   "Carrier_69_SpareSafetyInput(2_6)" AT %I3814.6 : Bool;   // SPARE SAFETY INPUT
   "Carrier_69_SpareSafetyInput(2_7)" AT %I3814.7 : Bool;   // SPARE SAFETY INPUT
   "Carrier_69_Slot3_SafetyOutput" AT %IW3815 : Word;   // SLOT 3 SAFETY OUTPUT WORD
   "Carrier_69_Crash_Detect_OK" AT %I3815.0 : Bool;   // CARRIER CRASH DETECT
   "Carrier_69_SpareSafetyOutput(3_1)" AT %I3815.1 : Bool;   // SPARE SAFETY OUTPUT
   "Carrier_69_SpareSafetyOutput(3_2)" AT %I3815.2 : Bool;   // SPARE SAFETY OUTPUT
   "Carrier_69_SpareSafetyOutput(3_3)" AT %I3815.3 : Bool;   // SPARE SAFETY OUTPUT
   "Carrier_69_SpareSafetyOutput(3_4)" AT %I3815.4 : Bool;   // SPARE SAFETY OUTPUT
   "Carrier_69_SpareSafetyOutput(3_5)" AT %I3815.5 : Bool;   // SPARE SAFETY OUTPUT
   "Carrier_69_SpareSafetyOutput(3_6)" AT %I3815.6 : Bool;   // SPARE SAFETY OUTPUT
   "Carrier_69_SpareSafetyOutput(3_7)" AT %I3815.7 : Bool;   // SPARE SAFETY OUTPUT
   "Carrier_69_Slot4_Input" AT %IW3816 : Word;   // SLOT 4 INPUT WORD
   "Carrier_69_480VPowerOn_MDCB1" AT %I3816.0 : Bool;   // 480 VAC POWER ON MDCB 1
   "Carrier_69_SpareInput(4_1)" AT %I3816.1 : Bool;   // SPARE INPUT
   "Carrier_69_SpareInput(4_2)" AT %I3816.2 : Bool;   // SPARE INPUT
   "Carrier_69_SitopSelectStatus" AT %I3816.3 : Bool;   // SITOP SELECT STATUS
   "Carrier_69_DCsupplyOnPSCB2" AT %I3816.4 : Bool;   // DC SUPPLY ON PSCB 2
   "Carrier_69_SpareInput(4_5)" AT %I3816.5 : Bool;   // SPARE INPUT
   "Carrier_69_SpareInput(4_6)" AT %I3816.6 : Bool;   // SPARE INPUT
   "Carrier_69_SpareInput(4_7)" AT %I3816.7 : Bool;   // SPARE INPUT
   "Carrier_69_PB1_ProdHoldLH" AT %I3817.0 : Bool;   // PB 1 PRODUCTION HOLD LH
   "Carrier_69_PB2_ResetLH" AT %I3817.1 : Bool;   // PB 2 RESET LH
   "Carrier_69_PB3_ProdHoldRH" AT %I3817.2 : Bool;   // PB 3 PRODUCTION HOLD RH
   "Carrier_69_PB4_ResetRH" AT %I3817.3 : Bool;   // PB 4 RESET RH
   "Carrier_69_SpareInput(4_14)" AT %I3817.4 : Bool;   // SPARE INPUT
   "Carrier_69_SpareInput(4_15)" AT %I3817.5 : Bool;   // SPARE INPUT
   "Carrier_69_SpareInput(4_16)" AT %I3817.6 : Bool;   // SPARE INPUT
   "Carrier_69_SpareInput(4_17)" AT %I3817.7 : Bool;   // SPARE INPUT
   "Carrier_69_Slot5_Output" AT %IW3818 : Word;   // SLOT 5 OUTPUT WORD
   "Carrier_69_IRD400_HMI_24VDC_ENABLE" AT %I3818.0 : Bool;   // IRD 400 PANEL HMI 24V DC POWER
   "Carrier_69_FaultLight_LH" AT %I3818.1 : Bool;   // FAULT LIGHT LH
   "Carrier_69_RunLight_LH" AT %I3818.2 : Bool;   // RUN LIGHT LH
   "Carrier_69_FaultLight_RH" AT %I3818.3 : Bool;   // FAULT LIGHT RH
   "Carrier_69_RunLight_RH" AT %I3818.4 : Bool;   // RUN LIGHT RH
   "Carrier_69_SpareOutput(5_5)" AT %I3818.5 : Bool;   // SPARE OUTPUT
   "Carrier_69_SpareOutput(5_6)" AT %I3818.6 : Bool;   // SPARE OUTPUT
   "Carrier_69_SpareOutput(5_7)" AT %I3818.7 : Bool;   // SPARE OUTPUT
   "Carrier_69_ActualSpeed" AT %IW3820 : Word;   // ACTUAL SPEED
   "Carrier_69_CarrierDriveAlarm" AT %IW3822 : Word;   // CARRIER DRIVE ALARM
   "Carrier_69_CarrierDriveWarning" AT %IW3824 : Word;   // CARRIER DRIVE WARNING
   "Carrier_70_Status" AT %IW3850 : Word;   // CARRIER STATUS WORD
   "Carrier_70_Status.0" AT %I3850.0 : Bool;   // HEARTBEAT
   "Carrier_70_Status.1" AT %I3850.1 : Bool;   // MANUAL
   "Carrier_70_Status.2" AT %I3850.2 : Bool;   // IN_AUTO
   "Carrier_70_Status.3" AT %I3850.3 : Bool;   // POSITIONING_COMPLETE
   "Carrier_70_Status.4" AT %I3850.4 : Bool;   // PRODUCTION HOLD
   "Carrier_70_Status.5" AT %I3850.5 : Bool;   // CARRIER MOVING FORWARD
   "Carrier_70_Status.6" AT %I3850.6 : Bool;   // CARRIER MOVING REVERSE
   "Carrier_70_Status.7" AT %I3850.7 : Bool;   // CARRIER FAULT
   "Carrier_70_Status.8" AT %I3851.0 : Bool;   // CRASH DETECT TRIPPED
   "Carrier_70_Status.9" AT %I3851.1 : Bool;
   "Carrier_70_Status.10" AT %I3851.2 : Bool;
   "Carrier_70_Status.11" AT %I3851.3 : Bool;
   "Carrier_70_Status.12" AT %I3851.4 : Bool;
   "Carrier_70_Status.13" AT %I3851.5 : Bool;
   "Carrier_70_Status.14" AT %I3851.6 : Bool;
   "Carrier_70_Status.15" AT %I3851.7 : Bool;
   "Carrier_70_SDCFaultCode" AT %IW3852 : Word;   // SDC FAULT CODE
   "Carrier_70_CarrierPosition" AT %ID3854 : DWord;   // CARRIER POSITION
   "Carrier_70_CarrierNumber" AT %IW3858 : Word;   // CARRIER NUMBER
   "Carrier_70_G120DControlWord" AT %IW3860 : Word;   // G120D_STW1_CONTROL
   "Carrier_70_G120DControlWord.0" AT %I3860.0 : Bool;   // Bit_00_ON
   "Carrier_70_G120DControlWord.1" AT %I3860.1 : Bool;   // Bit_01_AUS2_INH
   "Carrier_70_G120DControlWord.2" AT %I3860.2 : Bool;   // Bit_02_AUS3_STOP
   "Carrier_70_G120DControlWord.3" AT %I3860.3 : Bool;   // Bit_03_EN
   "Carrier_70_G120DControlWord.4" AT %I3860.4 : Bool;   // Bit_04_EN_RAMP
   "Carrier_70_G120DControlWord.5" AT %I3860.5 : Bool;   // Bit_05_START_RAMP
   "Carrier_70_G120DControlWord.6" AT %I3860.6 : Bool;   // Bit_06_SETPOINT
   "Carrier_70_G120DControlWord.7" AT %I3860.7 : Bool;   // Bit_07_RESET
   "Carrier_70_G120DControlWord.8" AT %I3861.0 : Bool;   // Bit_08_JOG_R
   "Carrier_70_G120DControlWord.9" AT %I3861.1 : Bool;   // Bit_09_JOG_L
   "Carrier_70_G120DControlWord.10" AT %I3861.2 : Bool;   // Bit_10_CONTR_PLC
   "Carrier_70_G120DControlWord.11" AT %I3861.3 : Bool;   // Bit_11_REVERSE
   "Carrier_70_G120DControlWord.12" AT %I3861.4 : Bool;   // Bit_12_BRAKE_RELEASE
   "Carrier_70_G120DControlWord.13" AT %I3861.5 : Bool;   // Bit_13_DDS
   "Carrier_70_G120DControlWord.14" AT %I3861.6 : Bool;   // Bit_14_DO0
   "Carrier_70_G120DControlWord.15" AT %I3861.7 : Bool;   // Bit_15_DO1
   "Carrier_70_G120DStatusWord" AT %IW3862 : Word;   // G120D_ZSW1_STATUS
   "Carrier_70_G120DStatusWord.0" AT %I3862.0 : Bool;   // Bit_00_READY_RUN
   "Carrier_70_G120DStatusWord.1" AT %I3862.1 : Bool;   // Bit_01_READY_ON
   "Carrier_70_G120DStatusWord.2" AT %I3862.2 : Bool;   // Bit_02_ENABLE
   "Carrier_70_G120DStatusWord.3" AT %I3862.3 : Bool;   // Bit_03_FAULT
   "Carrier_70_G120DStatusWord.4" AT %I3862.4 : Bool;   // Bit_04_OFF2
   "Carrier_70_G120DStatusWord.5" AT %I3862.5 : Bool;   // Bit_05_OFF3
   "Carrier_70_G120DStatusWord.6" AT %I3862.6 : Bool;   // Bit_06_LOCK_OUT
   "Carrier_70_G120DStatusWord.7" AT %I3862.7 : Bool;   // Bit_07_WARN
   "Carrier_70_G120DStatusWord.8" AT %I3863.0 : Bool;   // Bit_08_NO_DEVIATION
   "Carrier_70_G120DStatusWord.9" AT %I3863.1 : Bool;   // Bit_09_CONTR_PLC
   "Carrier_70_G120DStatusWord.10" AT %I3863.2 : Bool;   // Bit_10_F_MAX
   "Carrier_70_G120DStatusWord.11" AT %I3863.3 : Bool;   // Bit_11_LIMIT_REACHED
   "Carrier_70_G120DStatusWord.12" AT %I3863.4 : Bool;   // Bit_12_BRAKE_OPEN
   "Carrier_70_G120DStatusWord.13" AT %I3863.5 : Bool;   // Bit_13_NO_OVERTEMP
   "Carrier_70_G120DStatusWord.14" AT %I3863.6 : Bool;   // Bit_14_CW_CCW
   "Carrier_70_G120DStatusWord.15" AT %I3863.7 : Bool;   // Bit_15_OVERL
   "Carrier_70_Slot2_Input" AT %IW3864 : Word;   // SLOT 2 INPUT WORD
   "Carrier_70_CrashDetectSW" AT %I3864.0 : Bool;   // CRASH DETECT SW
   "Carrier_70_SpareSafetyInput(2_1)" AT %I3864.1 : Bool;   // SPARE SAFETY INPUT
   "Carrier_70_SpareSafetyInput(2_2)" AT %I3864.2 : Bool;   // SPARE SAFETY INPUT
   "Carrier_70_SpareSafetyInput(2_3)" AT %I3864.3 : Bool;   // SPARE SAFETY INPUT
   "Carrier_70_SpareSafetyInput(2_4)" AT %I3864.4 : Bool;   // SPARE SAFETY INPUT
   "Carrier_70_SpareSafetyInput(2_5)" AT %I3864.5 : Bool;   // SPARE SAFETY INPUT
   "Carrier_70_SpareSafetyInput(2_6)" AT %I3864.6 : Bool;   // SPARE SAFETY INPUT
   "Carrier_70_SpareSafetyInput(2_7)" AT %I3864.7 : Bool;   // SPARE SAFETY INPUT
   "Carrier_70_Slot3_SafetyOutput" AT %IW3865 : Word;   // SLOT 3 SAFETY OUTPUT WORD
   "Carrier_70_Crash_Detect_OK" AT %I3865.0 : Bool;   // CARRIER CRASH DETECT
   "Carrier_70_SpareSafetyOutput(3_1)" AT %I3865.1 : Bool;   // SPARE SAFETY OUTPUT
   "Carrier_70_SpareSafetyOutput(3_2)" AT %I3865.2 : Bool;   // SPARE SAFETY OUTPUT
   "Carrier_70_SpareSafetyOutput(3_3)" AT %I3865.3 : Bool;   // SPARE SAFETY OUTPUT
   "Carrier_70_SpareSafetyOutput(3_4)" AT %I3865.4 : Bool;   // SPARE SAFETY OUTPUT
   "Carrier_70_SpareSafetyOutput(3_5)" AT %I3865.5 : Bool;   // SPARE SAFETY OUTPUT
   "Carrier_70_SpareSafetyOutput(3_6)" AT %I3865.6 : Bool;   // SPARE SAFETY OUTPUT
   "Carrier_70_SpareSafetyOutput(3_7)" AT %I3865.7 : Bool;   // SPARE SAFETY OUTPUT
   "Carrier_70_Slot4_Input" AT %IW3866 : Word;   // SLOT 4 INPUT WORD
   "Carrier_70_480VPowerOn_MDCB1" AT %I3866.0 : Bool;   // 480 VAC POWER ON MDCB 1
   "Carrier_70_SpareInput(4_1)" AT %I3866.1 : Bool;   // SPARE INPUT
   "Carrier_70_SpareInput(4_2)" AT %I3866.2 : Bool;   // SPARE INPUT
   "Carrier_70_SitopSelectStatus" AT %I3866.3 : Bool;   // SITOP SELECT STATUS
   "Carrier_70_DCsupplyOnPSCB2" AT %I3866.4 : Bool;   // DC SUPPLY ON PSCB 2
   "Carrier_70_SpareInput(4_5)" AT %I3866.5 : Bool;   // SPARE INPUT
   "Carrier_70_SpareInput(4_6)" AT %I3866.6 : Bool;   // SPARE INPUT
   "Carrier_70_SpareInput(4_7)" AT %I3866.7 : Bool;   // SPARE INPUT
   "Carrier_70_PB1_ProdHoldLH" AT %I3867.0 : Bool;   // PB 1 PRODUCTION HOLD LH
   "Carrier_70_PB2_ResetLH" AT %I3867.1 : Bool;   // PB 2 RESET LH
   "Carrier_70_PB3_ProdHoldRH" AT %I3867.2 : Bool;   // PB 3 PRODUCTION HOLD RH
   "Carrier_70_PB4_ResetRH" AT %I3867.3 : Bool;   // PB 4 RESET RH
   "Carrier_70_SpareInput(4_14)" AT %I3867.4 : Bool;   // SPARE INPUT
   "Carrier_70_SpareInput(4_15)" AT %I3867.5 : Bool;   // SPARE INPUT
   "Carrier_70_SpareInput(4_16)" AT %I3867.6 : Bool;   // SPARE INPUT
   "Carrier_70_SpareInput(4_17)" AT %I3867.7 : Bool;   // SPARE INPUT
   "Carrier_70_Slot5_Output" AT %IW3868 : Word;   // SLOT 5 OUTPUT WORD
   "Carrier_70_IRD400_HMI_24VDC_ENABLE" AT %I3868.0 : Bool;   // IRD 400 PANEL HMI 24V DC POWER
   "Carrier_70_FaultLight_LH" AT %I3868.1 : Bool;   // FAULT LIGHT LH
   "Carrier_70_RunLight_LH" AT %I3868.2 : Bool;   // RUN LIGHT LH
   "Carrier_70_FaultLight_RH" AT %I3868.3 : Bool;   // FAULT LIGHT RH
   "Carrier_70_RunLight_RH" AT %I3868.4 : Bool;   // RUN LIGHT RH
   "Carrier_70_SpareOutput(5_5)" AT %I3868.5 : Bool;   // SPARE OUTPUT
   "Carrier_70_SpareOutput(5_6)" AT %I3868.6 : Bool;   // SPARE OUTPUT
   "Carrier_70_SpareOutput(5_7)" AT %I3868.7 : Bool;   // SPARE OUTPUT
   "Carrier_70_ActualSpeed" AT %IW3870 : Word;   // ACTUAL SPEED
   "Carrier_70_CarrierDriveAlarm" AT %IW3872 : Word;   // CARRIER DRIVE ALARM
   "Carrier_70_CarrierDriveWarning" AT %IW3874 : Word;   // CARRIER DRIVE WARNING
   "Carrier_71_Status" AT %IW3900 : Word;   // CARRIER STATUS WORD
   "Carrier_71_Status.0" AT %I3900.0 : Bool;   // HEARTBEAT
   "Carrier_71_Status.1" AT %I3900.1 : Bool;   // MANUAL
   "Carrier_71_Status.2" AT %I3900.2 : Bool;   // IN_AUTO
   "Carrier_71_Status.3" AT %I3900.3 : Bool;   // POSITIONING_COMPLETE
   "Carrier_71_Status.4" AT %I3900.4 : Bool;   // PRODUCTION HOLD
   "Carrier_71_Status.5" AT %I3900.5 : Bool;   // CARRIER MOVING FORWARD
   "Carrier_71_Status.6" AT %I3900.6 : Bool;   // CARRIER MOVING REVERSE
   "Carrier_71_Status.7" AT %I3900.7 : Bool;   // CARRIER FAULT
   "Carrier_71_Status.8" AT %I3901.0 : Bool;   // CRASH DETECT TRIPPED
   "Carrier_71_Status.9" AT %I3901.1 : Bool;
   "Carrier_71_Status.10" AT %I3901.2 : Bool;
   "Carrier_71_Status.11" AT %I3901.3 : Bool;
   "Carrier_71_Status.12" AT %I3901.4 : Bool;
   "Carrier_71_Status.13" AT %I3901.5 : Bool;
   "Carrier_71_Status.14" AT %I3901.6 : Bool;
   "Carrier_71_Status.15" AT %I3901.7 : Bool;
   "Carrier_71_SDCFaultCode" AT %IW3902 : Word;   // SDC FAULT CODE
   "Carrier_71_CarrierPosition" AT %ID3904 : DWord;   // CARRIER POSITION
   "Carrier_71_CarrierNumber" AT %IW3908 : Word;   // CARRIER NUMBER
   "Carrier_71_G120DControlWord" AT %IW3910 : Word;   // G120D_STW1_CONTROL
   "Carrier_71_G120DControlWord.0" AT %I3910.0 : Bool;   // Bit_00_ON
   "Carrier_71_G120DControlWord.1" AT %I3910.1 : Bool;   // Bit_01_AUS2_INH
   "Carrier_71_G120DControlWord.2" AT %I3910.2 : Bool;   // Bit_02_AUS3_STOP
   "Carrier_71_G120DControlWord.3" AT %I3910.3 : Bool;   // Bit_03_EN
   "Carrier_71_G120DControlWord.4" AT %I3910.4 : Bool;   // Bit_04_EN_RAMP
   "Carrier_71_G120DControlWord.5" AT %I3910.5 : Bool;   // Bit_05_START_RAMP
   "Carrier_71_G120DControlWord.6" AT %I3910.6 : Bool;   // Bit_06_SETPOINT
   "Carrier_71_G120DControlWord.7" AT %I3910.7 : Bool;   // Bit_07_RESET
   "Carrier_71_G120DControlWord.8" AT %I3911.0 : Bool;   // Bit_08_JOG_R
   "Carrier_71_G120DControlWord.9" AT %I3911.1 : Bool;   // Bit_09_JOG_L
   "Carrier_71_G120DControlWord.10" AT %I3911.2 : Bool;   // Bit_10_CONTR_PLC
   "Carrier_71_G120DControlWord.11" AT %I3911.3 : Bool;   // Bit_11_REVERSE
   "Carrier_71_G120DControlWord.12" AT %I3911.4 : Bool;   // Bit_12_BRAKE_RELEASE
   "Carrier_71_G120DControlWord.13" AT %I3911.5 : Bool;   // Bit_13_DDS
   "Carrier_71_G120DControlWord.14" AT %I3911.6 : Bool;   // Bit_14_DO0
   "Carrier_71_G120DControlWord.15" AT %I3911.7 : Bool;   // Bit_15_DO1
   "Carrier_71_G120DStatusWord" AT %IW3912 : Word;   // G120D_ZSW1_STATUS
   "Carrier_71_G120DStatusWord.0" AT %I3912.0 : Bool;   // Bit_00_READY_RUN
   "Carrier_71_G120DStatusWord.1" AT %I3912.1 : Bool;   // Bit_01_READY_ON
   "Carrier_71_G120DStatusWord.2" AT %I3912.2 : Bool;   // Bit_02_ENABLE
   "Carrier_71_G120DStatusWord.3" AT %I3912.3 : Bool;   // Bit_03_FAULT
   "Carrier_71_G120DStatusWord.4" AT %I3912.4 : Bool;   // Bit_04_OFF2
   "Carrier_71_G120DStatusWord.5" AT %I3912.5 : Bool;   // Bit_05_OFF3
   "Carrier_71_G120DStatusWord.6" AT %I3912.6 : Bool;   // Bit_06_LOCK_OUT
   "Carrier_71_G120DStatusWord.7" AT %I3912.7 : Bool;   // Bit_07_WARN
   "Carrier_71_G120DStatusWord.8" AT %I3913.0 : Bool;   // Bit_08_NO_DEVIATION
   "Carrier_71_G120DStatusWord.9" AT %I3913.1 : Bool;   // Bit_09_CONTR_PLC
   "Carrier_71_G120DStatusWord.10" AT %I3913.2 : Bool;   // Bit_10_F_MAX
   "Carrier_71_G120DStatusWord.11" AT %I3913.3 : Bool;   // Bit_11_LIMIT_REACHED
   "Carrier_71_G120DStatusWord.12" AT %I3913.4 : Bool;   // Bit_12_BRAKE_OPEN
   "Carrier_71_G120DStatusWord.13" AT %I3913.5 : Bool;   // Bit_13_NO_OVERTEMP
   "Carrier_71_G120DStatusWord.14" AT %I3913.6 : Bool;   // Bit_14_CW_CCW
   "Carrier_71_G120DStatusWord.15" AT %I3913.7 : Bool;   // Bit_15_OVERL
   "Carrier_71_Slot2_Input" AT %IW3914 : Word;   // SLOT 2 INPUT WORD
   "Carrier_71_CrashDetectSW" AT %I3914.0 : Bool;   // CRASH DETECT SW
   "Carrier_71_SpareSafetyInput(2_1)" AT %I3914.1 : Bool;   // SPARE SAFETY INPUT
   "Carrier_71_SpareSafetyInput(2_2)" AT %I3914.2 : Bool;   // SPARE SAFETY INPUT
   "Carrier_71_SpareSafetyInput(2_3)" AT %I3914.3 : Bool;   // SPARE SAFETY INPUT
   "Carrier_71_SpareSafetyInput(2_4)" AT %I3914.4 : Bool;   // SPARE SAFETY INPUT
   "Carrier_71_SpareSafetyInput(2_5)" AT %I3914.5 : Bool;   // SPARE SAFETY INPUT
   "Carrier_71_SpareSafetyInput(2_6)" AT %I3914.6 : Bool;   // SPARE SAFETY INPUT
   "Carrier_71_SpareSafetyInput(2_7)" AT %I3914.7 : Bool;   // SPARE SAFETY INPUT
   "Carrier_71_Slot3_SafetyOutput" AT %IW3915 : Word;   // SLOT 3 SAFETY OUTPUT WORD
   "Carrier_71_Crash_Detect_OK" AT %I3915.0 : Bool;   // CARRIER CRASH DETECT
   "Carrier_71_SpareSafetyOutput(3_1)" AT %I3915.1 : Bool;   // SPARE SAFETY OUTPUT
   "Carrier_71_SpareSafetyOutput(3_2)" AT %I3915.2 : Bool;   // SPARE SAFETY OUTPUT
   "Carrier_71_SpareSafetyOutput(3_3)" AT %I3915.3 : Bool;   // SPARE SAFETY OUTPUT
   "Carrier_71_SpareSafetyOutput(3_4)" AT %I3915.4 : Bool;   // SPARE SAFETY OUTPUT
   "Carrier_71_SpareSafetyOutput(3_5)" AT %I3915.5 : Bool;   // SPARE SAFETY OUTPUT
   "Carrier_71_SpareSafetyOutput(3_6)" AT %I3915.6 : Bool;   // SPARE SAFETY OUTPUT
   "Carrier_71_SpareSafetyOutput(3_7)" AT %I3915.7 : Bool;   // SPARE SAFETY OUTPUT
   "Carrier_71_Slot4_Input" AT %IW3916 : Word;   // SLOT 4 INPUT WORD
   "Carrier_71_480VPowerOn_MDCB1" AT %I3916.0 : Bool;   // 480 VAC POWER ON MDCB 1
   "Carrier_71_SpareInput(4_1)" AT %I3916.1 : Bool;   // SPARE INPUT
   "Carrier_71_SpareInput(4_2)" AT %I3916.2 : Bool;   // SPARE INPUT
   "Carrier_71_SitopSelectStatus" AT %I3916.3 : Bool;   // SITOP SELECT STATUS
   "Carrier_71_DCsupplyOnPSCB2" AT %I3916.4 : Bool;   // DC SUPPLY ON PSCB 2
   "Carrier_71_SpareInput(4_5)" AT %I3916.5 : Bool;   // SPARE INPUT
   "Carrier_71_SpareInput(4_6)" AT %I3916.6 : Bool;   // SPARE INPUT
   "Carrier_71_SpareInput(4_7)" AT %I3916.7 : Bool;   // SPARE INPUT
   "Carrier_71_PB1_ProdHoldLH" AT %I3917.0 : Bool;   // PB 1 PRODUCTION HOLD LH
   "Carrier_71_PB2_ResetLH" AT %I3917.1 : Bool;   // PB 2 RESET LH
   "Carrier_71_PB3_ProdHoldRH" AT %I3917.2 : Bool;   // PB 3 PRODUCTION HOLD RH
   "Carrier_71_PB4_ResetRH" AT %I3917.3 : Bool;   // PB 4 RESET RH
   "Carrier_71_SpareInput(4_14)" AT %I3917.4 : Bool;   // SPARE INPUT
   "Carrier_71_SpareInput(4_15)" AT %I3917.5 : Bool;   // SPARE INPUT
   "Carrier_71_SpareInput(4_16)" AT %I3917.6 : Bool;   // SPARE INPUT
   "Carrier_71_SpareInput(4_17)" AT %I3917.7 : Bool;   // SPARE INPUT
   "Carrier_71_Slot5_Output" AT %IW3918 : Word;   // SLOT 5 OUTPUT WORD
   "Carrier_71_IRD400_HMI_24VDC_ENABLE" AT %I3918.0 : Bool;   // IRD 400 PANEL HMI 24V DC POWER
   "Carrier_71_FaultLight_LH" AT %I3918.1 : Bool;   // FAULT LIGHT LH
   "Carrier_71_RunLight_LH" AT %I3918.2 : Bool;   // RUN LIGHT LH
   "Carrier_71_FaultLight_RH" AT %I3918.3 : Bool;   // FAULT LIGHT RH
   "Carrier_71_RunLight_RH" AT %I3918.4 : Bool;   // RUN LIGHT RH
   "Carrier_71_SpareOutput(5_5)" AT %I3918.5 : Bool;   // SPARE OUTPUT
   "Carrier_71_SpareOutput(5_6)" AT %I3918.6 : Bool;   // SPARE OUTPUT
   "Carrier_71_SpareOutput(5_7)" AT %I3918.7 : Bool;   // SPARE OUTPUT
   "Carrier_71_ActualSpeed" AT %IW3920 : Word;   // ACTUAL SPEED
   "Carrier_71_CarrierDriveAlarm" AT %IW3922 : Word;   // CARRIER DRIVE ALARM
   "Carrier_71_CarrierDriveWarning" AT %IW3924 : Word;   // CARRIER DRIVE WARNING
   "Carrier_72_Status" AT %IW3950 : Word;   // CARRIER STATUS WORD
   "Carrier_72_Status.0" AT %I3950.0 : Bool;   // HEARTBEAT
   "Carrier_72_Status.1" AT %I3950.1 : Bool;   // MANUAL
   "Carrier_72_Status.2" AT %I3950.2 : Bool;   // IN_AUTO
   "Carrier_72_Status.3" AT %I3950.3 : Bool;   // POSITIONING_COMPLETE
   "Carrier_72_Status.4" AT %I3950.4 : Bool;   // PRODUCTION HOLD
   "Carrier_72_Status.5" AT %I3950.5 : Bool;   // CARRIER MOVING FORWARD
   "Carrier_72_Status.6" AT %I3950.6 : Bool;   // CARRIER MOVING REVERSE
   "Carrier_72_Status.7" AT %I3950.7 : Bool;   // CARRIER FAULT
   "Carrier_72_Status.8" AT %I3951.0 : Bool;   // CRASH DETECT TRIPPED
   "Carrier_72_Status.9" AT %I3951.1 : Bool;
   "Carrier_72_Status.10" AT %I3951.2 : Bool;
   "Carrier_72_Status.11" AT %I3951.3 : Bool;
   "Carrier_72_Status.12" AT %I3951.4 : Bool;
   "Carrier_72_Status.13" AT %I3951.5 : Bool;
   "Carrier_72_Status.14" AT %I3951.6 : Bool;
   "Carrier_72_Status.15" AT %I3951.7 : Bool;
   "Carrier_72_SDCFaultCode" AT %IW3952 : Word;   // SDC FAULT CODE
   "Carrier_72_CarrierPosition" AT %ID3954 : DWord;   // CARRIER POSITION
   "Carrier_72_CarrierNumber" AT %IW3958 : Word;   // CARRIER NUMBER
   "Carrier_72_G120DControlWord" AT %IW3960 : Word;   // G120D_STW1_CONTROL
   "Carrier_72_G120DControlWord.0" AT %I3960.0 : Bool;   // Bit_00_ON
   "Carrier_72_G120DControlWord.1" AT %I3960.1 : Bool;   // Bit_01_AUS2_INH
   "Carrier_72_G120DControlWord.2" AT %I3960.2 : Bool;   // Bit_02_AUS3_STOP
   "Carrier_72_G120DControlWord.3" AT %I3960.3 : Bool;   // Bit_03_EN
   "Carrier_72_G120DControlWord.4" AT %I3960.4 : Bool;   // Bit_04_EN_RAMP
   "Carrier_72_G120DControlWord.5" AT %I3960.5 : Bool;   // Bit_05_START_RAMP
   "Carrier_72_G120DControlWord.6" AT %I3960.6 : Bool;   // Bit_06_SETPOINT
   "Carrier_72_G120DControlWord.7" AT %I3960.7 : Bool;   // Bit_07_RESET
   "Carrier_72_G120DControlWord.8" AT %I3961.0 : Bool;   // Bit_08_JOG_R
   "Carrier_72_G120DControlWord.9" AT %I3961.1 : Bool;   // Bit_09_JOG_L
   "Carrier_72_G120DControlWord.10" AT %I3961.2 : Bool;   // Bit_10_CONTR_PLC
   "Carrier_72_G120DControlWord.11" AT %I3961.3 : Bool;   // Bit_11_REVERSE
   "Carrier_72_G120DControlWord.12" AT %I3961.4 : Bool;   // Bit_12_BRAKE_RELEASE
   "Carrier_72_G120DControlWord.13" AT %I3961.5 : Bool;   // Bit_13_DDS
   "Carrier_72_G120DControlWord.14" AT %I3961.6 : Bool;   // Bit_14_DO0
   "Carrier_72_G120DControlWord.15" AT %I3961.7 : Bool;   // Bit_15_DO1
   "Carrier_72_G120DStatusWord" AT %IW3962 : Word;   // G120D_ZSW1_STATUS
   "Carrier_72_G120DStatusWord.0" AT %I3962.0 : Bool;   // Bit_00_READY_RUN
   "Carrier_72_G120DStatusWord.1" AT %I3962.1 : Bool;   // Bit_01_READY_ON
   "Carrier_72_G120DStatusWord.2" AT %I3962.2 : Bool;   // Bit_02_ENABLE
   "Carrier_72_G120DStatusWord.3" AT %I3962.3 : Bool;   // Bit_03_FAULT
   "Carrier_72_G120DStatusWord.4" AT %I3962.4 : Bool;   // Bit_04_OFF2
   "Carrier_72_G120DStatusWord.5" AT %I3962.5 : Bool;   // Bit_05_OFF3
   "Carrier_72_G120DStatusWord.6" AT %I3962.6 : Bool;   // Bit_06_LOCK_OUT
   "Carrier_72_G120DStatusWord.7" AT %I3962.7 : Bool;   // Bit_07_WARN
   "Carrier_72_G120DStatusWord.8" AT %I3963.0 : Bool;   // Bit_08_NO_DEVIATION
   "Carrier_72_G120DStatusWord.9" AT %I3963.1 : Bool;   // Bit_09_CONTR_PLC
   "Carrier_72_G120DStatusWord.10" AT %I3963.2 : Bool;   // Bit_10_F_MAX
   "Carrier_72_G120DStatusWord.11" AT %I3963.3 : Bool;   // Bit_11_LIMIT_REACHED
   "Carrier_72_G120DStatusWord.12" AT %I3963.4 : Bool;   // Bit_12_BRAKE_OPEN
   "Carrier_72_G120DStatusWord.13" AT %I3963.5 : Bool;   // Bit_13_NO_OVERTEMP
   "Carrier_72_G120DStatusWord.14" AT %I3963.6 : Bool;   // Bit_14_CW_CCW
   "Carrier_72_G120DStatusWord.15" AT %I3963.7 : Bool;   // Bit_15_OVERL
   "Carrier_72_Slot2_Input" AT %IW3964 : Word;   // SLOT 2 INPUT WORD
   "Carrier_72_CrashDetectSW" AT %I3964.0 : Bool;   // CRASH DETECT SW
   "Carrier_72_SpareSafetyInput(2_1)" AT %I3964.1 : Bool;   // SPARE SAFETY INPUT
   "Carrier_72_SpareSafetyInput(2_2)" AT %I3964.2 : Bool;   // SPARE SAFETY INPUT
   "Carrier_72_SpareSafetyInput(2_3)" AT %I3964.3 : Bool;   // SPARE SAFETY INPUT
   "Carrier_72_SpareSafetyInput(2_4)" AT %I3964.4 : Bool;   // SPARE SAFETY INPUT
   "Carrier_72_SpareSafetyInput(2_5)" AT %I3964.5 : Bool;   // SPARE SAFETY INPUT
   "Carrier_72_SpareSafetyInput(2_6)" AT %I3964.6 : Bool;   // SPARE SAFETY INPUT
   "Carrier_72_SpareSafetyInput(2_7)" AT %I3964.7 : Bool;   // SPARE SAFETY INPUT
   "Carrier_72_Slot3_SafetyOutput" AT %IW3965 : Word;   // SLOT 3 SAFETY OUTPUT WORD
   "Carrier_72_Crash_Detect_OK" AT %I3965.0 : Bool;   // CARRIER CRASH DETECT
   "Carrier_72_SpareSafetyOutput(3_1)" AT %I3965.1 : Bool;   // SPARE SAFETY OUTPUT
   "Carrier_72_SpareSafetyOutput(3_2)" AT %I3965.2 : Bool;   // SPARE SAFETY OUTPUT
   "Carrier_72_SpareSafetyOutput(3_3)" AT %I3965.3 : Bool;   // SPARE SAFETY OUTPUT
   "Carrier_72_SpareSafetyOutput(3_4)" AT %I3965.4 : Bool;   // SPARE SAFETY OUTPUT
   "Carrier_72_SpareSafetyOutput(3_5)" AT %I3965.5 : Bool;   // SPARE SAFETY OUTPUT
   "Carrier_72_SpareSafetyOutput(3_6)" AT %I3965.6 : Bool;   // SPARE SAFETY OUTPUT
   "Carrier_72_SpareSafetyOutput(3_7)" AT %I3965.7 : Bool;   // SPARE SAFETY OUTPUT
   "Carrier_72_Slot4_Input" AT %IW3966 : Word;   // SLOT 4 INPUT WORD
   "Carrier_72_480VPowerOn_MDCB1" AT %I3966.0 : Bool;   // 480 VAC POWER ON MDCB 1
   "Carrier_72_SpareInput(4_1)" AT %I3966.1 : Bool;   // SPARE INPUT
   "Carrier_72_SpareInput(4_2)" AT %I3966.2 : Bool;   // SPARE INPUT
   "Carrier_72_SitopSelectStatus" AT %I3966.3 : Bool;   // SITOP SELECT STATUS
   "Carrier_72_DCsupplyOnPSCB2" AT %I3966.4 : Bool;   // DC SUPPLY ON PSCB 2
   "Carrier_72_SpareInput(4_5)" AT %I3966.5 : Bool;   // SPARE INPUT
   "Carrier_72_SpareInput(4_6)" AT %I3966.6 : Bool;   // SPARE INPUT
   "Carrier_72_SpareInput(4_7)" AT %I3966.7 : Bool;   // SPARE INPUT
   "Carrier_72_PB1_ProdHoldLH" AT %I3967.0 : Bool;   // PB 1 PRODUCTION HOLD LH
   "Carrier_72_PB2_ResetLH" AT %I3967.1 : Bool;   // PB 2 RESET LH
   "Carrier_72_PB3_ProdHoldRH" AT %I3967.2 : Bool;   // PB 3 PRODUCTION HOLD RH
   "Carrier_72_PB4_ResetRH" AT %I3967.3 : Bool;   // PB 4 RESET RH
   "Carrier_72_SpareInput(4_14)" AT %I3967.4 : Bool;   // SPARE INPUT
   "Carrier_72_SpareInput(4_15)" AT %I3967.5 : Bool;   // SPARE INPUT
   "Carrier_72_SpareInput(4_16)" AT %I3967.6 : Bool;   // SPARE INPUT
   "Carrier_72_SpareInput(4_17)" AT %I3967.7 : Bool;   // SPARE INPUT
   "Carrier_72_Slot5_Output" AT %IW3968 : Word;   // SLOT 5 OUTPUT WORD
   "Carrier_72_IRD400_HMI_24VDC_ENABLE" AT %I3968.0 : Bool;   // IRD 400 PANEL HMI 24V DC POWER
   "Carrier_72_FaultLight_LH" AT %I3968.1 : Bool;   // FAULT LIGHT LH
   "Carrier_72_RunLight_LH" AT %I3968.2 : Bool;   // RUN LIGHT LH
   "Carrier_72_FaultLight_RH" AT %I3968.3 : Bool;   // FAULT LIGHT RH
   "Carrier_72_RunLight_RH" AT %I3968.4 : Bool;   // RUN LIGHT RH
   "Carrier_72_SpareOutput(5_5)" AT %I3968.5 : Bool;   // SPARE OUTPUT
   "Carrier_72_SpareOutput(5_6)" AT %I3968.6 : Bool;   // SPARE OUTPUT
   "Carrier_72_SpareOutput(5_7)" AT %I3968.7 : Bool;   // SPARE OUTPUT
   "Carrier_72_ActualSpeed" AT %IW3970 : Word;   // ACTUAL SPEED
   "Carrier_72_CarrierDriveAlarm" AT %IW3972 : Word;   // CARRIER DRIVE ALARM
   "Carrier_72_CarrierDriveWarning" AT %IW3974 : Word;   // CARRIER DRIVE WARNING
   "Carrier_73_Status" AT %IW4000 : Word;   // CARRIER STATUS WORD
   "Carrier_73_Status.0" AT %I4000.0 : Bool;   // HEARTBEAT
   "Carrier_73_Status.1" AT %I4000.1 : Bool;   // MANUAL
   "Carrier_73_Status.2" AT %I4000.2 : Bool;   // IN_AUTO
   "Carrier_73_Status.3" AT %I4000.3 : Bool;   // POSITIONING_COMPLETE
   "Carrier_73_Status.4" AT %I4000.4 : Bool;   // PRODUCTION HOLD
   "Carrier_73_Status.5" AT %I4000.5 : Bool;   // CARRIER MOVING FORWARD
   "Carrier_73_Status.6" AT %I4000.6 : Bool;   // CARRIER MOVING REVERSE
   "Carrier_73_Status.7" AT %I4000.7 : Bool;   // CARRIER FAULT
   "Carrier_73_Status.8" AT %I4001.0 : Bool;   // CRASH DETECT TRIPPED
   "Carrier_73_Status.9" AT %I4001.1 : Bool;
   "Carrier_73_Status.10" AT %I4001.2 : Bool;
   "Carrier_73_Status.11" AT %I4001.3 : Bool;
   "Carrier_73_Status.12" AT %I4001.4 : Bool;
   "Carrier_73_Status.13" AT %I4001.5 : Bool;
   "Carrier_73_Status.14" AT %I4001.6 : Bool;
   "Carrier_73_Status.15" AT %I4001.7 : Bool;
   "Carrier_73_SDCFaultCode" AT %IW4002 : Word;   // SDC FAULT CODE
   "Carrier_73_CarrierPosition" AT %ID4004 : DWord;   // CARRIER POSITION
   "Carrier_73_CarrierNumber" AT %IW4008 : Word;   // CARRIER NUMBER
   "Carrier_73_G120DControlWord" AT %IW4010 : Word;   // G120D_STW1_CONTROL
   "Carrier_73_G120DControlWord.0" AT %I4010.0 : Bool;   // Bit_00_ON
   "Carrier_73_G120DControlWord.1" AT %I4010.1 : Bool;   // Bit_01_AUS2_INH
   "Carrier_73_G120DControlWord.2" AT %I4010.2 : Bool;   // Bit_02_AUS3_STOP
   "Carrier_73_G120DControlWord.3" AT %I4010.3 : Bool;   // Bit_03_EN
   "Carrier_73_G120DControlWord.4" AT %I4010.4 : Bool;   // Bit_04_EN_RAMP
   "Carrier_73_G120DControlWord.5" AT %I4010.5 : Bool;   // Bit_05_START_RAMP
   "Carrier_73_G120DControlWord.6" AT %I4010.6 : Bool;   // Bit_06_SETPOINT
   "Carrier_73_G120DControlWord.7" AT %I4010.7 : Bool;   // Bit_07_RESET
   "Carrier_73_G120DControlWord.8" AT %I4011.0 : Bool;   // Bit_08_JOG_R
   "Carrier_73_G120DControlWord.9" AT %I4011.1 : Bool;   // Bit_09_JOG_L
   "Carrier_73_G120DControlWord.10" AT %I4011.2 : Bool;   // Bit_10_CONTR_PLC
   "Carrier_73_G120DControlWord.11" AT %I4011.3 : Bool;   // Bit_11_REVERSE
   "Carrier_73_G120DControlWord.12" AT %I4011.4 : Bool;   // Bit_12_BRAKE_RELEASE
   "Carrier_73_G120DControlWord.13" AT %I4011.5 : Bool;   // Bit_13_DDS
   "Carrier_73_G120DControlWord.14" AT %I4011.6 : Bool;   // Bit_14_DO0
   "Carrier_73_G120DControlWord.15" AT %I4011.7 : Bool;   // Bit_15_DO1
   "Carrier_73_G120DStatusWord" AT %IW4012 : Word;   // G120D_ZSW1_STATUS
   "Carrier_73_G120DStatusWord.0" AT %I4012.0 : Bool;   // Bit_00_READY_RUN
   "Carrier_73_G120DStatusWord.1" AT %I4012.1 : Bool;   // Bit_01_READY_ON
   "Carrier_73_G120DStatusWord.2" AT %I4012.2 : Bool;   // Bit_02_ENABLE
   "Carrier_73_G120DStatusWord.3" AT %I4012.3 : Bool;   // Bit_03_FAULT
   "Carrier_73_G120DStatusWord.4" AT %I4012.4 : Bool;   // Bit_04_OFF2
   "Carrier_73_G120DStatusWord.5" AT %I4012.5 : Bool;   // Bit_05_OFF3
   "Carrier_73_G120DStatusWord.6" AT %I4012.6 : Bool;   // Bit_06_LOCK_OUT
   "Carrier_73_G120DStatusWord.7" AT %I4012.7 : Bool;   // Bit_07_WARN
   "Carrier_73_G120DStatusWord.8" AT %I4013.0 : Bool;   // Bit_08_NO_DEVIATION
   "Carrier_73_G120DStatusWord.9" AT %I4013.1 : Bool;   // Bit_09_CONTR_PLC
   "Carrier_73_G120DStatusWord.10" AT %I4013.2 : Bool;   // Bit_10_F_MAX
   "Carrier_73_G120DStatusWord.11" AT %I4013.3 : Bool;   // Bit_11_LIMIT_REACHED
   "Carrier_73_G120DStatusWord.12" AT %I4013.4 : Bool;   // Bit_12_BRAKE_OPEN
   "Carrier_73_G120DStatusWord.13" AT %I4013.5 : Bool;   // Bit_13_NO_OVERTEMP
   "Carrier_73_G120DStatusWord.14" AT %I4013.6 : Bool;   // Bit_14_CW_CCW
   "Carrier_73_G120DStatusWord.15" AT %I4013.7 : Bool;   // Bit_15_OVERL
   "Carrier_73_Slot2_Input" AT %IW4014 : Word;   // SLOT 2 INPUT WORD
   "Carrier_73_CrashDetectSW" AT %I4014.0 : Bool;   // CRASH DETECT SW
   "Carrier_73_SpareSafetyInput(2_1)" AT %I4014.1 : Bool;   // SPARE SAFETY INPUT
   "Carrier_73_SpareSafetyInput(2_2)" AT %I4014.2 : Bool;   // SPARE SAFETY INPUT
   "Carrier_73_SpareSafetyInput(2_3)" AT %I4014.3 : Bool;   // SPARE SAFETY INPUT
   "Carrier_73_SpareSafetyInput(2_4)" AT %I4014.4 : Bool;   // SPARE SAFETY INPUT
   "Carrier_73_SpareSafetyInput(2_5)" AT %I4014.5 : Bool;   // SPARE SAFETY INPUT
   "Carrier_73_SpareSafetyInput(2_6)" AT %I4014.6 : Bool;   // SPARE SAFETY INPUT
   "Carrier_73_SpareSafetyInput(2_7)" AT %I4014.7 : Bool;   // SPARE SAFETY INPUT
   "Carrier_73_Slot3_SafetyOutput" AT %IW4015 : Word;   // SLOT 3 SAFETY OUTPUT WORD
   "Carrier_73_Crash_Detect_OK" AT %I4015.0 : Bool;   // CARRIER CRASH DETECT
   "Carrier_73_SpareSafetyOutput(3_1)" AT %I4015.1 : Bool;   // SPARE SAFETY OUTPUT
   "Carrier_73_SpareSafetyOutput(3_2)" AT %I4015.2 : Bool;   // SPARE SAFETY OUTPUT
   "Carrier_73_SpareSafetyOutput(3_3)" AT %I4015.3 : Bool;   // SPARE SAFETY OUTPUT
   "Carrier_73_SpareSafetyOutput(3_4)" AT %I4015.4 : Bool;   // SPARE SAFETY OUTPUT
   "Carrier_73_SpareSafetyOutput(3_5)" AT %I4015.5 : Bool;   // SPARE SAFETY OUTPUT
   "Carrier_73_SpareSafetyOutput(3_6)" AT %I4015.6 : Bool;   // SPARE SAFETY OUTPUT
   "Carrier_73_SpareSafetyOutput(3_7)" AT %I4015.7 : Bool;   // SPARE SAFETY OUTPUT
   "Carrier_73_Slot4_Input" AT %IW4016 : Word;   // SLOT 4 INPUT WORD
   "Carrier_73_480VPowerOn_MDCB1" AT %I4016.0 : Bool;   // 480 VAC POWER ON MDCB 1
   "Carrier_73_SpareInput(4_1)" AT %I4016.1 : Bool;   // SPARE INPUT
   "Carrier_73_SpareInput(4_2)" AT %I4016.2 : Bool;   // SPARE INPUT
   "Carrier_73_SitopSelectStatus" AT %I4016.3 : Bool;   // SITOP SELECT STATUS
   "Carrier_73_DCsupplyOnPSCB2" AT %I4016.4 : Bool;   // DC SUPPLY ON PSCB 2
   "Carrier_73_SpareInput(4_5)" AT %I4016.5 : Bool;   // SPARE INPUT
   "Carrier_73_SpareInput(4_6)" AT %I4016.6 : Bool;   // SPARE INPUT
   "Carrier_73_SpareInput(4_7)" AT %I4016.7 : Bool;   // SPARE INPUT
   "Carrier_73_PB1_ProdHoldLH" AT %I4017.0 : Bool;   // PB 1 PRODUCTION HOLD LH
   "Carrier_73_PB2_ResetLH" AT %I4017.1 : Bool;   // PB 2 RESET LH
   "Carrier_73_PB3_ProdHoldRH" AT %I4017.2 : Bool;   // PB 3 PRODUCTION HOLD RH
   "Carrier_73_PB4_ResetRH" AT %I4017.3 : Bool;   // PB 4 RESET RH
   "Carrier_73_SpareInput(4_14)" AT %I4017.4 : Bool;   // SPARE INPUT
   "Carrier_73_SpareInput(4_15)" AT %I4017.5 : Bool;   // SPARE INPUT
   "Carrier_73_SpareInput(4_16)" AT %I4017.6 : Bool;   // SPARE INPUT
   "Carrier_73_SpareInput(4_17)" AT %I4017.7 : Bool;   // SPARE INPUT
   "Carrier_73_Slot5_Output" AT %IW4018 : Word;   // SLOT 5 OUTPUT WORD
   "Carrier_73_IRD400_HMI_24VDC_ENABLE" AT %I4018.0 : Bool;   // IRD 400 PANEL HMI 24V DC POWER
   "Carrier_73_FaultLight_LH" AT %I4018.1 : Bool;   // FAULT LIGHT LH
   "Carrier_73_RunLight_LH" AT %I4018.2 : Bool;   // RUN LIGHT LH
   "Carrier_73_FaultLight_RH" AT %I4018.3 : Bool;   // FAULT LIGHT RH
   "Carrier_73_RunLight_RH" AT %I4018.4 : Bool;   // RUN LIGHT RH
   "Carrier_73_SpareOutput(5_5)" AT %I4018.5 : Bool;   // SPARE OUTPUT
   "Carrier_73_SpareOutput(5_6)" AT %I4018.6 : Bool;   // SPARE OUTPUT
   "Carrier_73_SpareOutput(5_7)" AT %I4018.7 : Bool;   // SPARE OUTPUT
   "Carrier_73_ActualSpeed" AT %IW4020 : Word;   // ACTUAL SPEED
   "Carrier_73_CarrierDriveAlarm" AT %IW4022 : Word;   // CARRIER DRIVE ALARM
   "Carrier_73_CarrierDriveWarning" AT %IW4024 : Word;   // CARRIER DRIVE WARNING
   "Carrier_74_Status" AT %IW4050 : Word;   // CARRIER STATUS WORD
   "Carrier_74_Status.0" AT %I4050.0 : Bool;   // HEARTBEAT
   "Carrier_74_Status.1" AT %I4050.1 : Bool;   // MANUAL
   "Carrier_74_Status.2" AT %I4050.2 : Bool;   // IN_AUTO
   "Carrier_74_Status.3" AT %I4050.3 : Bool;   // POSITIONING_COMPLETE
   "Carrier_74_Status.4" AT %I4050.4 : Bool;   // PRODUCTION HOLD
   "Carrier_74_Status.5" AT %I4050.5 : Bool;   // CARRIER MOVING FORWARD
   "Carrier_74_Status.6" AT %I4050.6 : Bool;   // CARRIER MOVING REVERSE